(* Logix 5000 project; controller FV vendor 1 type 14 code 217 rev 31.11; software revision 31.00; part 38 of 63 *)
(* tags used below, declared in another part *)
   CWD : CHECKWORD_FLAGS;
   Dummy : BOOL;
   FV_Copy_from_fv_file : DINT;
   FV_Copy_to_fv_file : DINT;
   FV_LTX_YS_001 : PlantItem;   // LTX_YS_001
   FV_LTX_YS_001_RawInput : ALIAS FOR Remote_IO:7:I.Data.16;   // FV_LTX_YS_001
   FV_LTX_YS_002 : PlantItem;   // LTX_YS_002
   FV_LTX_YS_002_RawInput : ALIAS FOR Remote_IO:7:I.Data.17;   // FV_LTX_YS_002
   FV_N110 : INT[255];   // FV DATA 0 CURRENT FV DATA
   FV_N111 : INT[50];   // FV1, CURRENT FV DATA
   FV_N112 : INT[50];   // FV2, CURRENT FV DATA
   FV_N113 : INT[50];   // FV3, CURRENT FV DATA
   FV_N114 : INT[50];   // FV4, CURRENT FV DATA
   FV_N115 : INT[50];   // FV5, CURRENT FV DATA
   FV_N116 : INT[50];   // FV6, CURRENT FV DATA
   FV_N117 : INT[50];   // FV7, CURRENT FV DATA
   FV_N118 : INT[50];   // FV8, CURRENT FV DATA
   FV_N119 : INT[50];   // FV9, CURRENT FV DATA
   FV_N120 : INT[50];   // FV10, CURRENT FV DATA
   FV_N121 : INT[50];   // FV11, CURRENT FV DATA
   FV_N122 : INT[50];   // FV12, CURRENT FV DATA
   FV_N123 : INT[50];   // FV13, CURRENT FV DATA
   FV_N124 : INT[50];   // FV14, CURRENT FV DATA
   FV_N125 : INT[50];   // FV15, CURRENT FV DATA
   FV_N126 : INT[50];   // FV16, CURRENT FV DATA
   FV_N127 : INT[50];   // FV17, CURRENT FV DATA
   FV_N128 : INT[50];   // FV18, CURRENT FV DATA
   FV_N129 : INT[50];   // FV19, CURRENT FV DATA
   FV_N130 : INT[50];   // FV20, CURRENT FV DATA
   FV_N131 : INT[50];   // FV21, CURRENT FV DATA
   FV_N132 : INT[50];   // FV22, CURRENT FV DATA
   FV_N133 : INT[50];   // FV23, CURRENT FV DATA
   FV_N134 : INT[50];   // FV24, CURRENT FV DATA
   FV_N135 : INT[50];   // FV25, CURRENT FV DATA
   FV_N136 : INT[50];   // YSV1, CURRENT FV DATA
   FV_N137 : INT[50];   // YSV2, CURRENT FV DATA
   FV_N138 : INT[50];   // YSV3, CURRENT FV DATA
   FV_N139 : INT[255];   // YST1
   FV_N140 : INT[255];   // YST2
   FV_N141 : INT[255];   // YSV1 DATA
   FV_N142 : INT[255];   // YSV2 DATA
   FV_N143 : INT[255];   // YSV3 DATA
   FV_N144 : INT[255];   // YST1 DATA
   FV_N145 : INT[255];   // YST2 DATA
   FV_N146 : INT[50];   // FV26, CURRENT FV DATA
   FV_N147 : INT[50];   // FV27, CURRENT FV DATA
   FV_N148 : INT[50];   // FV28, CURRENT FV DATA
   FV_N149 : INT[50];   // FV29, CURRENT FV DATA
   FV_N150 : INT[50];   // FV30, CURRENT FV DATA
   FV_N151 : INT[50];   // FV31, CURRENT FV DATA
   FV_PX1 : PlantItem;   // PX1
   FV_PX1_RawInput : ALIAS FOR Remote_IO:6:I.Data.13;   // FV_PX1 Water flush proxy switch
   FV_PX2 : PlantItem;   // PX2
   FV_PX2_RawInput : ALIAS FOR Remote_IO:6:I.Data.14;   // FV_PX2 CIP supply proxy switch
   FV_PX3 : PlantItem;   // PX3
   FV_PX3_RawInput : ALIAS FOR Remote_IO:6:I.Data.15;   // FV_PX3 YSV1 to reseeding main proxy switch
   One_Second_One_Scan : ALIAS FOR One_Second_1_scan;
(* FV_Common, continued *)

ROUTINE FV_Copy_Vessel_File   (* ladder *)
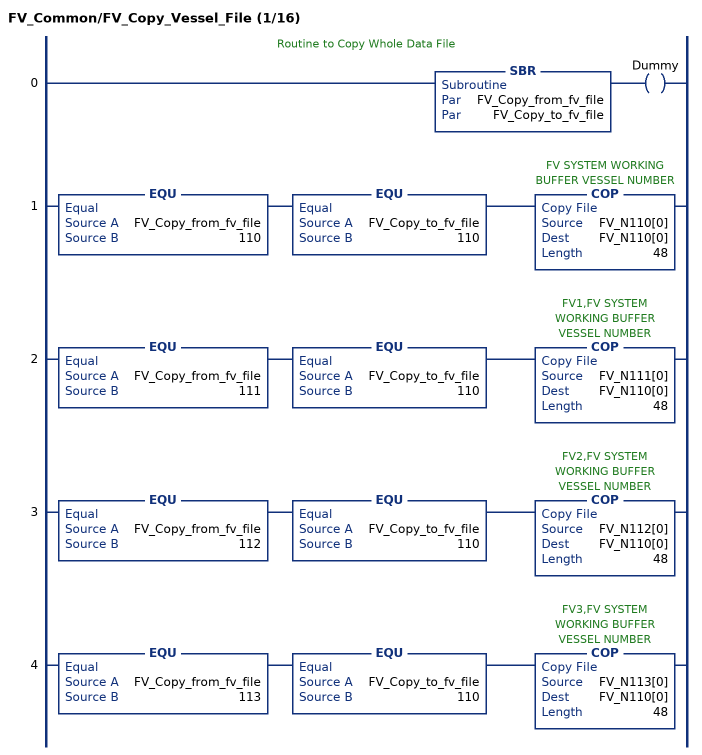
   // Routine to Copy Whole Data File
   0: SBR(FV_Copy_from_fv_file,FV_Copy_to_fv_file)OTE(Dummy);
   1: EQU(FV_Copy_from_fv_file,110)EQU(FV_Copy_to_fv_file,110)COP(FV_N110[0],FV_N110[0],48);
   2: EQU(FV_Copy_from_fv_file,111)EQU(FV_Copy_to_fv_file,110)COP(FV_N111[0],FV_N110[0],48);
   3: EQU(FV_Copy_from_fv_file,112)EQU(FV_Copy_to_fv_file,110)COP(FV_N112[0],FV_N110[0],48);
   4: EQU(FV_Copy_from_fv_file,113)EQU(FV_Copy_to_fv_file,110)COP(FV_N113[0],FV_N110[0],48);
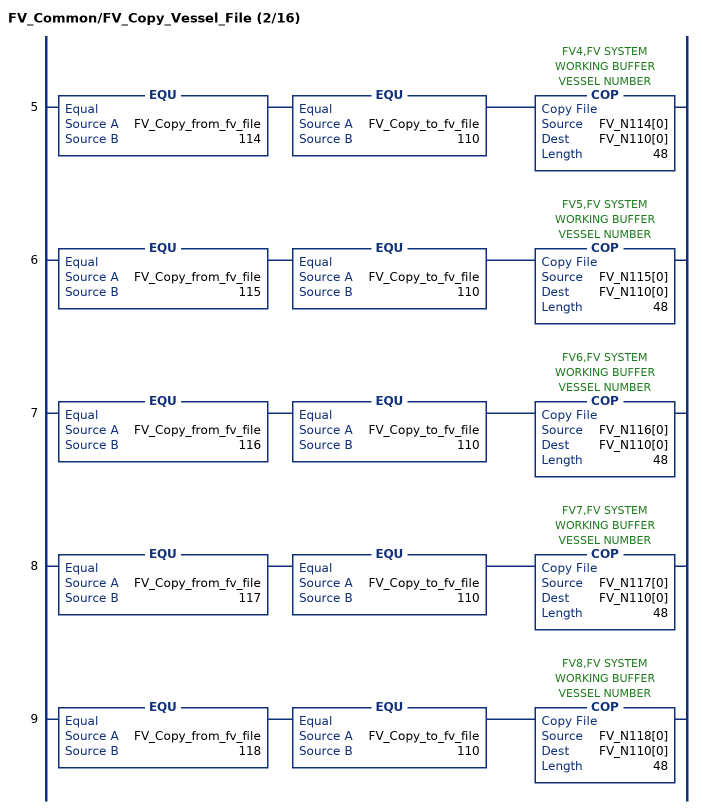
   5: EQU(FV_Copy_from_fv_file,114)EQU(FV_Copy_to_fv_file,110)COP(FV_N114[0],FV_N110[0],48);
   6: EQU(FV_Copy_from_fv_file,115)EQU(FV_Copy_to_fv_file,110)COP(FV_N115[0],FV_N110[0],48);
   7: EQU(FV_Copy_from_fv_file,116)EQU(FV_Copy_to_fv_file,110)COP(FV_N116[0],FV_N110[0],48);
   8: EQU(FV_Copy_from_fv_file,117)EQU(FV_Copy_to_fv_file,110)COP(FV_N117[0],FV_N110[0],48);
   9: EQU(FV_Copy_from_fv_file,118)EQU(FV_Copy_to_fv_file,110)COP(FV_N118[0],FV_N110[0],48);
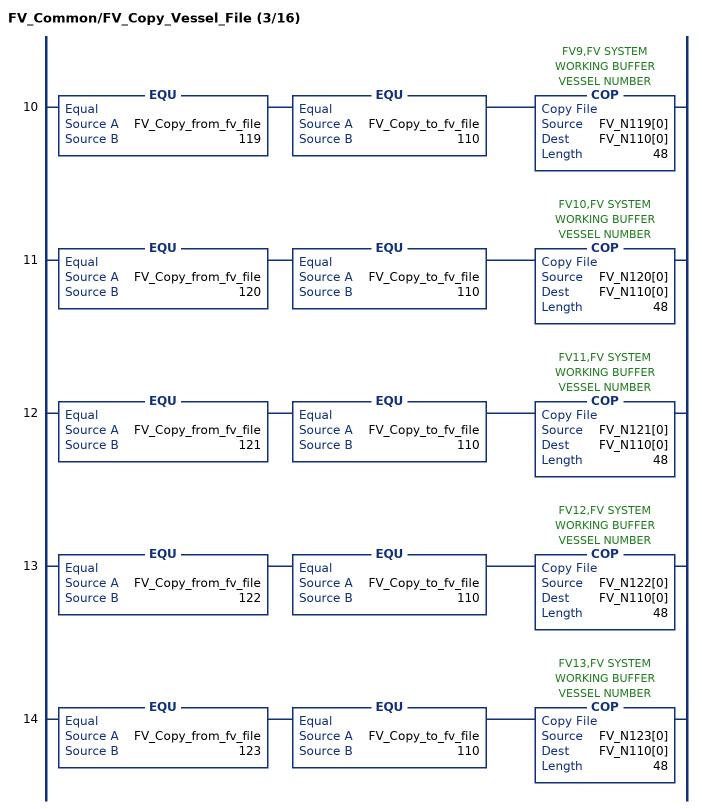
   10: EQU(FV_Copy_from_fv_file,119)EQU(FV_Copy_to_fv_file,110)COP(FV_N119[0],FV_N110[0],48);
   11: EQU(FV_Copy_from_fv_file,120)EQU(FV_Copy_to_fv_file,110)COP(FV_N120[0],FV_N110[0],48);
   12: EQU(FV_Copy_from_fv_file,121)EQU(FV_Copy_to_fv_file,110)COP(FV_N121[0],FV_N110[0],48);
   13: EQU(FV_Copy_from_fv_file,122)EQU(FV_Copy_to_fv_file,110)COP(FV_N122[0],FV_N110[0],48);
   14: EQU(FV_Copy_from_fv_file,123)EQU(FV_Copy_to_fv_file,110)COP(FV_N123[0],FV_N110[0],48);
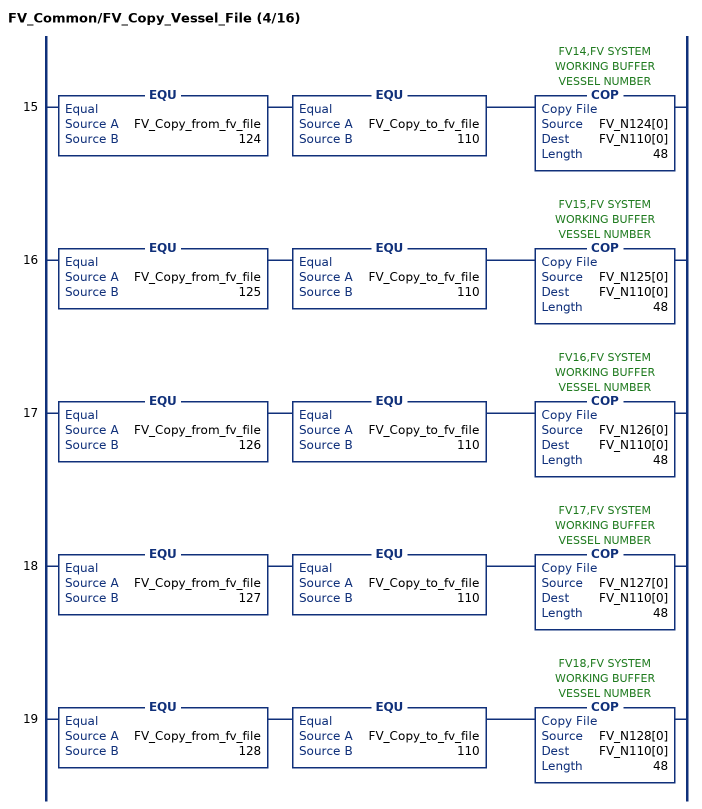
   15: EQU(FV_Copy_from_fv_file,124)EQU(FV_Copy_to_fv_file,110)COP(FV_N124[0],FV_N110[0],48);
   16: EQU(FV_Copy_from_fv_file,125)EQU(FV_Copy_to_fv_file,110)COP(FV_N125[0],FV_N110[0],48);
   17: EQU(FV_Copy_from_fv_file,126)EQU(FV_Copy_to_fv_file,110)COP(FV_N126[0],FV_N110[0],48);
   18: EQU(FV_Copy_from_fv_file,127)EQU(FV_Copy_to_fv_file,110)COP(FV_N127[0],FV_N110[0],48);
   19: EQU(FV_Copy_from_fv_file,128)EQU(FV_Copy_to_fv_file,110)COP(FV_N128[0],FV_N110[0],48);
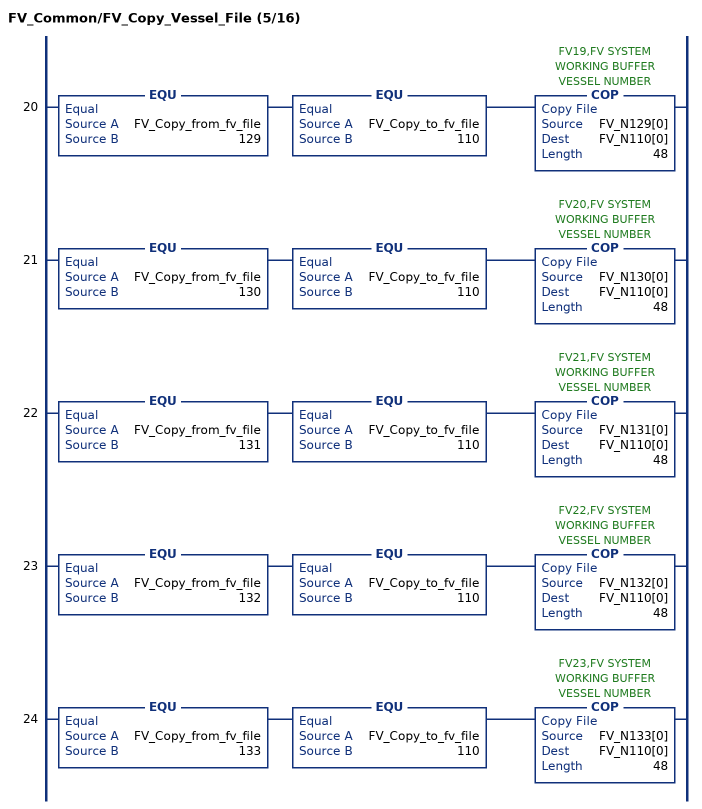
   20: EQU(FV_Copy_from_fv_file,129)EQU(FV_Copy_to_fv_file,110)COP(FV_N129[0],FV_N110[0],48);
   21: EQU(FV_Copy_from_fv_file,130)EQU(FV_Copy_to_fv_file,110)COP(FV_N130[0],FV_N110[0],48);
   22: EQU(FV_Copy_from_fv_file,131)EQU(FV_Copy_to_fv_file,110)COP(FV_N131[0],FV_N110[0],48);
   23: EQU(FV_Copy_from_fv_file,132)EQU(FV_Copy_to_fv_file,110)COP(FV_N132[0],FV_N110[0],48);
   24: EQU(FV_Copy_from_fv_file,133)EQU(FV_Copy_to_fv_file,110)COP(FV_N133[0],FV_N110[0],48);
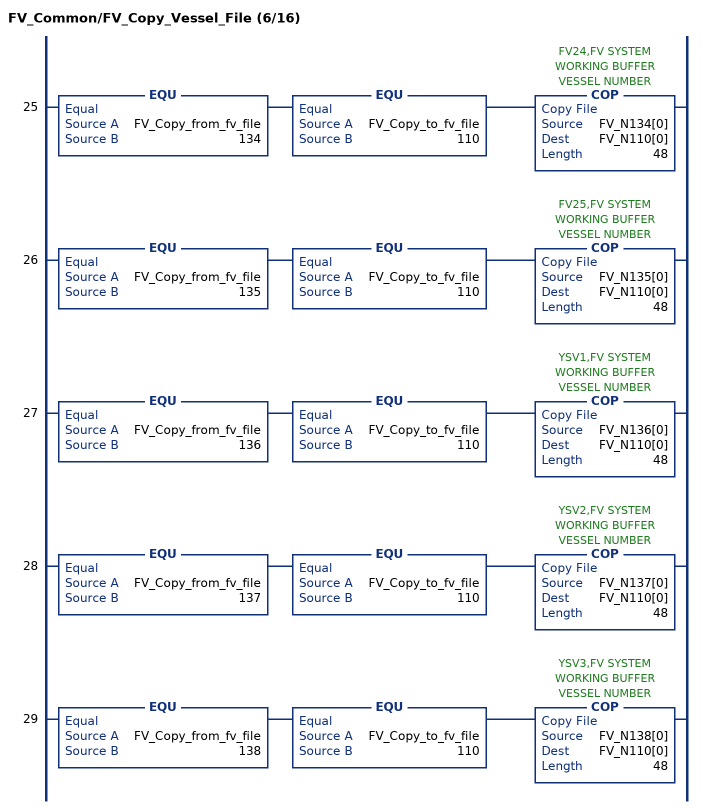
   25: EQU(FV_Copy_from_fv_file,134)EQU(FV_Copy_to_fv_file,110)COP(FV_N134[0],FV_N110[0],48);
   26: EQU(FV_Copy_from_fv_file,135)EQU(FV_Copy_to_fv_file,110)COP(FV_N135[0],FV_N110[0],48);
   27: EQU(FV_Copy_from_fv_file,136)EQU(FV_Copy_to_fv_file,110)COP(FV_N136[0],FV_N110[0],48);
   28: EQU(FV_Copy_from_fv_file,137)EQU(FV_Copy_to_fv_file,110)COP(FV_N137[0],FV_N110[0],48);
   29: EQU(FV_Copy_from_fv_file,138)EQU(FV_Copy_to_fv_file,110)COP(FV_N138[0],FV_N110[0],48);
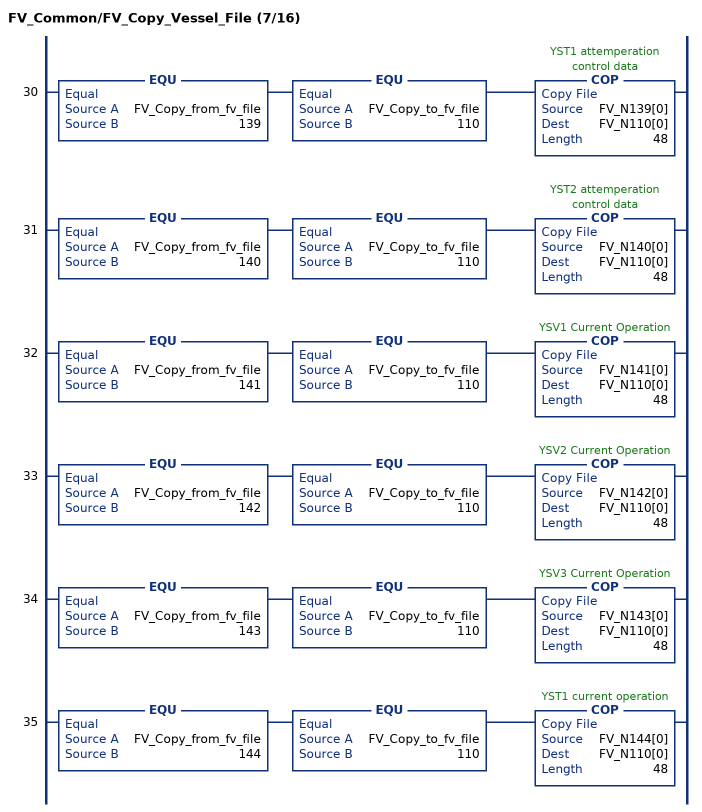
   30: EQU(FV_Copy_from_fv_file,139)EQU(FV_Copy_to_fv_file,110)COP(FV_N139[0],FV_N110[0],48);
   31: EQU(FV_Copy_from_fv_file,140)EQU(FV_Copy_to_fv_file,110)COP(FV_N140[0],FV_N110[0],48);
   32: EQU(FV_Copy_from_fv_file,141)EQU(FV_Copy_to_fv_file,110)COP(FV_N141[0],FV_N110[0],48);
   33: EQU(FV_Copy_from_fv_file,142)EQU(FV_Copy_to_fv_file,110)COP(FV_N142[0],FV_N110[0],48);
   34: EQU(FV_Copy_from_fv_file,143)EQU(FV_Copy_to_fv_file,110)COP(FV_N143[0],FV_N110[0],48);
   35: EQU(FV_Copy_from_fv_file,144)EQU(FV_Copy_to_fv_file,110)COP(FV_N144[0],FV_N110[0],48);
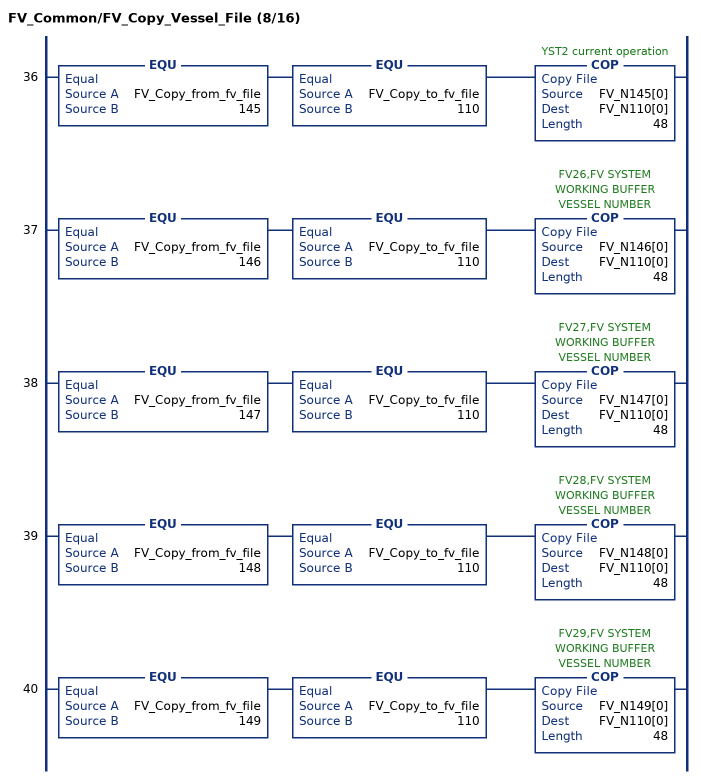
   36: EQU(FV_Copy_from_fv_file,145)EQU(FV_Copy_to_fv_file,110)COP(FV_N145[0],FV_N110[0],48);
   37: EQU(FV_Copy_from_fv_file,146)EQU(FV_Copy_to_fv_file,110)COP(FV_N146[0],FV_N110[0],48);
   38: EQU(FV_Copy_from_fv_file,147)EQU(FV_Copy_to_fv_file,110)COP(FV_N147[0],FV_N110[0],48);
   39: EQU(FV_Copy_from_fv_file,148)EQU(FV_Copy_to_fv_file,110)COP(FV_N148[0],FV_N110[0],48);
   40: EQU(FV_Copy_from_fv_file,149)EQU(FV_Copy_to_fv_file,110)COP(FV_N149[0],FV_N110[0],48);
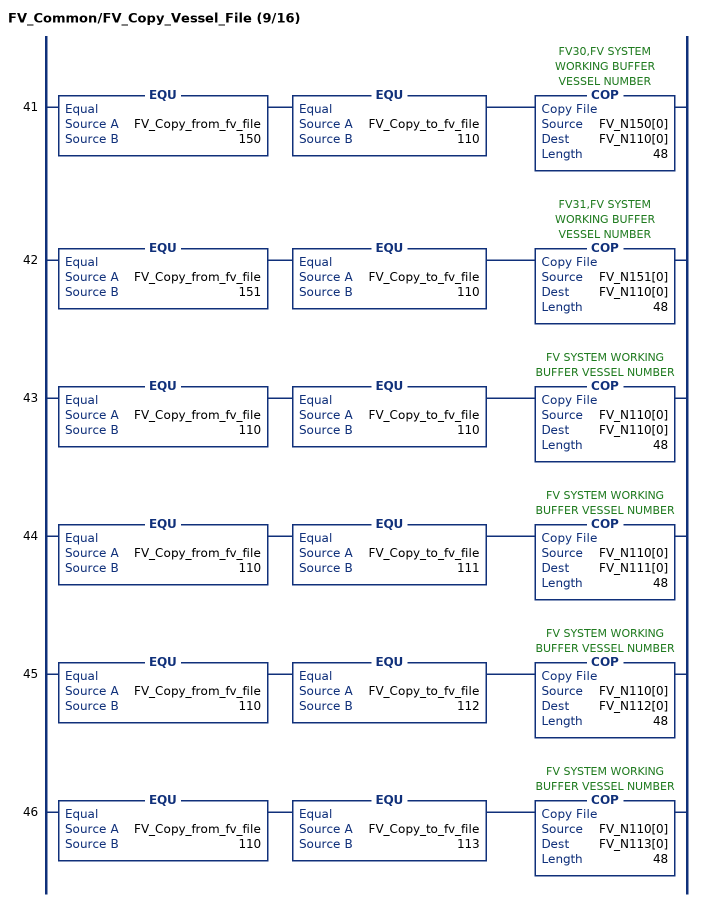
   41: EQU(FV_Copy_from_fv_file,150)EQU(FV_Copy_to_fv_file,110)COP(FV_N150[0],FV_N110[0],48);
   42: EQU(FV_Copy_from_fv_file,151)EQU(FV_Copy_to_fv_file,110)COP(FV_N151[0],FV_N110[0],48);
   43: EQU(FV_Copy_from_fv_file,110)EQU(FV_Copy_to_fv_file,110)COP(FV_N110[0],FV_N110[0],48);
   44: EQU(FV_Copy_from_fv_file,110)EQU(FV_Copy_to_fv_file,111)COP(FV_N110[0],FV_N111[0],48);
   45: EQU(FV_Copy_from_fv_file,110)EQU(FV_Copy_to_fv_file,112)COP(FV_N110[0],FV_N112[0],48);
   46: EQU(FV_Copy_from_fv_file,110)EQU(FV_Copy_to_fv_file,113)COP(FV_N110[0],FV_N113[0],48);
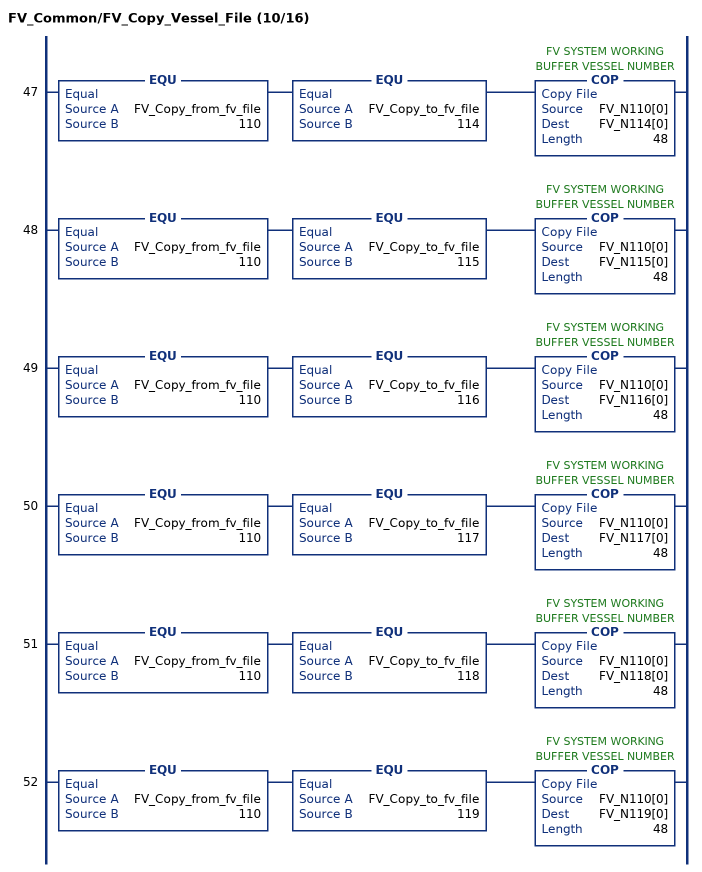
   47: EQU(FV_Copy_from_fv_file,110)EQU(FV_Copy_to_fv_file,114)COP(FV_N110[0],FV_N114[0],48);
   48: EQU(FV_Copy_from_fv_file,110)EQU(FV_Copy_to_fv_file,115)COP(FV_N110[0],FV_N115[0],48);
   49: EQU(FV_Copy_from_fv_file,110)EQU(FV_Copy_to_fv_file,116)COP(FV_N110[0],FV_N116[0],48);
   50: EQU(FV_Copy_from_fv_file,110)EQU(FV_Copy_to_fv_file,117)COP(FV_N110[0],FV_N117[0],48);
   51: EQU(FV_Copy_from_fv_file,110)EQU(FV_Copy_to_fv_file,118)COP(FV_N110[0],FV_N118[0],48);
   52: EQU(FV_Copy_from_fv_file,110)EQU(FV_Copy_to_fv_file,119)COP(FV_N110[0],FV_N119[0],48);
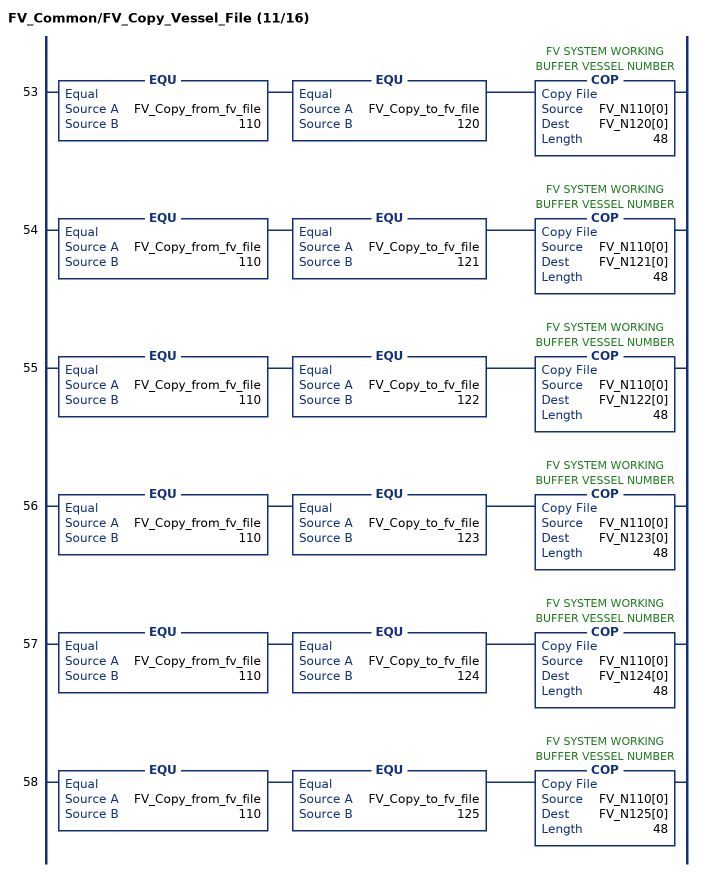
   53: EQU(FV_Copy_from_fv_file,110)EQU(FV_Copy_to_fv_file,120)COP(FV_N110[0],FV_N120[0],48);
   54: EQU(FV_Copy_from_fv_file,110)EQU(FV_Copy_to_fv_file,121)COP(FV_N110[0],FV_N121[0],48);
   55: EQU(FV_Copy_from_fv_file,110)EQU(FV_Copy_to_fv_file,122)COP(FV_N110[0],FV_N122[0],48);
   56: EQU(FV_Copy_from_fv_file,110)EQU(FV_Copy_to_fv_file,123)COP(FV_N110[0],FV_N123[0],48);
   57: EQU(FV_Copy_from_fv_file,110)EQU(FV_Copy_to_fv_file,124)COP(FV_N110[0],FV_N124[0],48);
   58: EQU(FV_Copy_from_fv_file,110)EQU(FV_Copy_to_fv_file,125)COP(FV_N110[0],FV_N125[0],48);
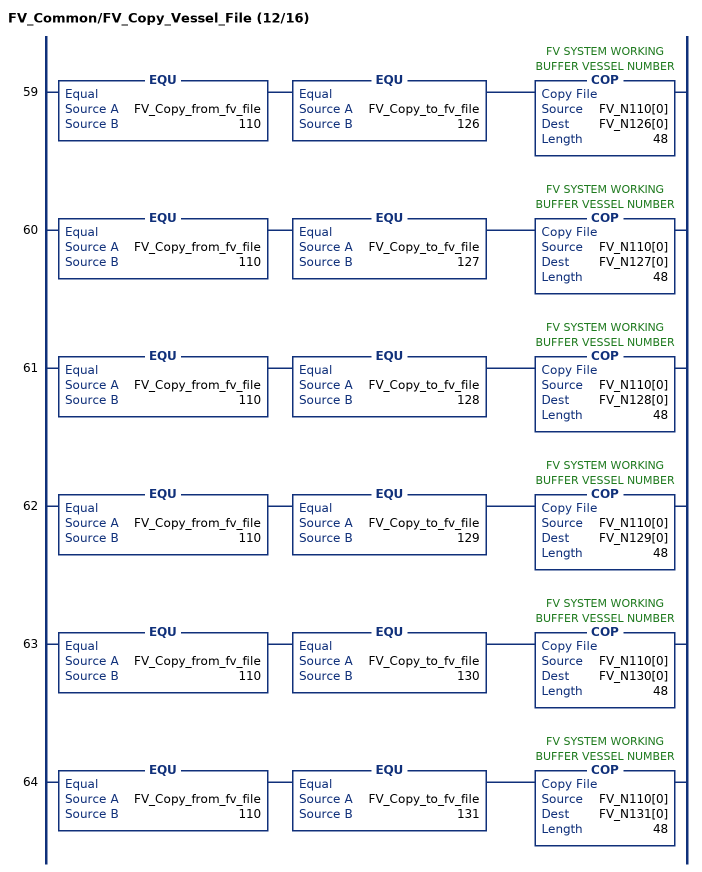
   59: EQU(FV_Copy_from_fv_file,110)EQU(FV_Copy_to_fv_file,126)COP(FV_N110[0],FV_N126[0],48);
   60: EQU(FV_Copy_from_fv_file,110)EQU(FV_Copy_to_fv_file,127)COP(FV_N110[0],FV_N127[0],48);
   61: EQU(FV_Copy_from_fv_file,110)EQU(FV_Copy_to_fv_file,128)COP(FV_N110[0],FV_N128[0],48);
   62: EQU(FV_Copy_from_fv_file,110)EQU(FV_Copy_to_fv_file,129)COP(FV_N110[0],FV_N129[0],48);
   63: EQU(FV_Copy_from_fv_file,110)EQU(FV_Copy_to_fv_file,130)COP(FV_N110[0],FV_N130[0],48);
   64: EQU(FV_Copy_from_fv_file,110)EQU(FV_Copy_to_fv_file,131)COP(FV_N110[0],FV_N131[0],48);
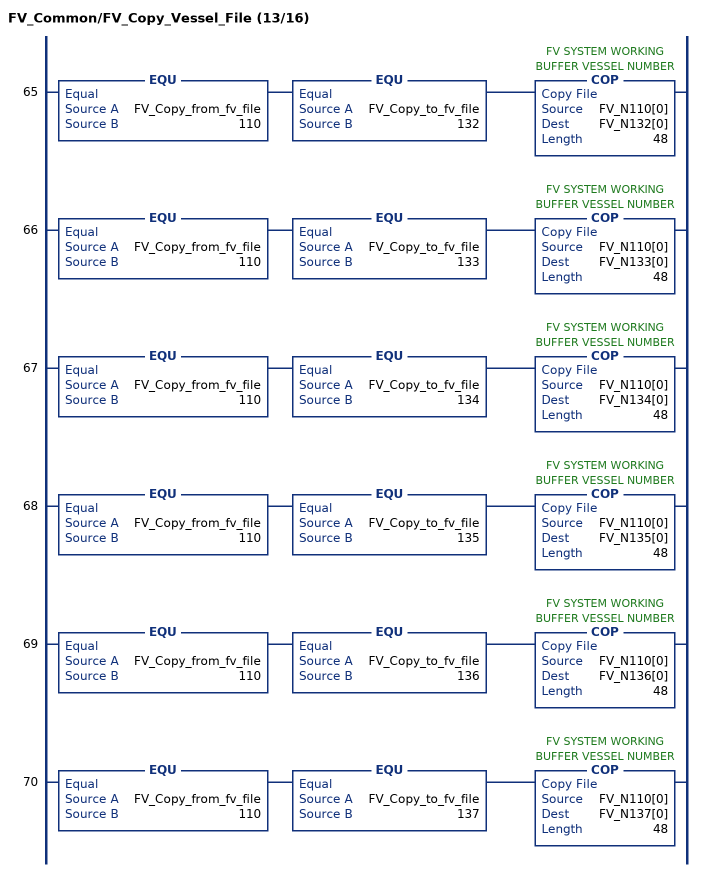
   65: EQU(FV_Copy_from_fv_file,110)EQU(FV_Copy_to_fv_file,132)COP(FV_N110[0],FV_N132[0],48);
   66: EQU(FV_Copy_from_fv_file,110)EQU(FV_Copy_to_fv_file,133)COP(FV_N110[0],FV_N133[0],48);
   67: EQU(FV_Copy_from_fv_file,110)EQU(FV_Copy_to_fv_file,134)COP(FV_N110[0],FV_N134[0],48);
   68: EQU(FV_Copy_from_fv_file,110)EQU(FV_Copy_to_fv_file,135)COP(FV_N110[0],FV_N135[0],48);
   69: EQU(FV_Copy_from_fv_file,110)EQU(FV_Copy_to_fv_file,136)COP(FV_N110[0],FV_N136[0],48);
   70: EQU(FV_Copy_from_fv_file,110)EQU(FV_Copy_to_fv_file,137)COP(FV_N110[0],FV_N137[0],48);
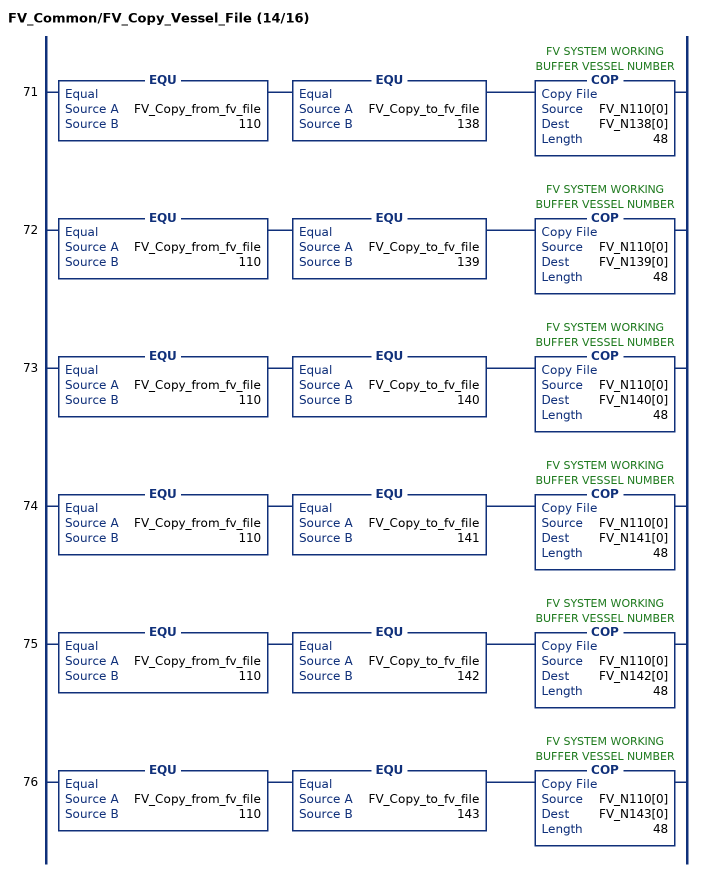
   71: EQU(FV_Copy_from_fv_file,110)EQU(FV_Copy_to_fv_file,138)COP(FV_N110[0],FV_N138[0],48);
   72: EQU(FV_Copy_from_fv_file,110)EQU(FV_Copy_to_fv_file,139)COP(FV_N110[0],FV_N139[0],48);
   73: EQU(FV_Copy_from_fv_file,110)EQU(FV_Copy_to_fv_file,140)COP(FV_N110[0],FV_N140[0],48);
   74: EQU(FV_Copy_from_fv_file,110)EQU(FV_Copy_to_fv_file,141)COP(FV_N110[0],FV_N141[0],48);
   75: EQU(FV_Copy_from_fv_file,110)EQU(FV_Copy_to_fv_file,142)COP(FV_N110[0],FV_N142[0],48);
   76: EQU(FV_Copy_from_fv_file,110)EQU(FV_Copy_to_fv_file,143)COP(FV_N110[0],FV_N143[0],48);
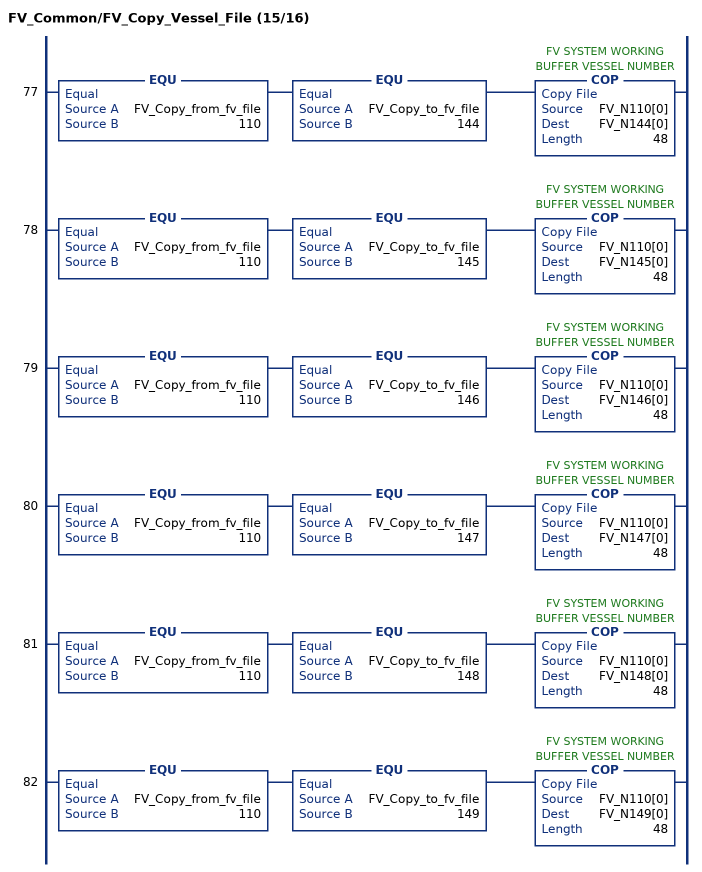
   77: EQU(FV_Copy_from_fv_file,110)EQU(FV_Copy_to_fv_file,144)COP(FV_N110[0],FV_N144[0],48);
   78: EQU(FV_Copy_from_fv_file,110)EQU(FV_Copy_to_fv_file,145)COP(FV_N110[0],FV_N145[0],48);
   79: EQU(FV_Copy_from_fv_file,110)EQU(FV_Copy_to_fv_file,146)COP(FV_N110[0],FV_N146[0],48);
   80: EQU(FV_Copy_from_fv_file,110)EQU(FV_Copy_to_fv_file,147)COP(FV_N110[0],FV_N147[0],48);
   81: EQU(FV_Copy_from_fv_file,110)EQU(FV_Copy_to_fv_file,148)COP(FV_N110[0],FV_N148[0],48);
   82: EQU(FV_Copy_from_fv_file,110)EQU(FV_Copy_to_fv_file,149)COP(FV_N110[0],FV_N149[0],48);
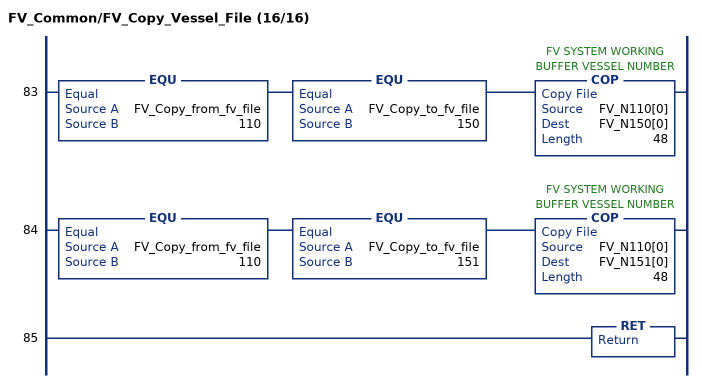
   83: EQU(FV_Copy_from_fv_file,110)EQU(FV_Copy_to_fv_file,150)COP(FV_N110[0],FV_N150[0],48);
   84: EQU(FV_Copy_from_fv_file,110)EQU(FV_Copy_to_fv_file,151)COP(FV_N110[0],FV_N151[0],48);
   85: RET();
END_ROUTINE

ROUTINE FV_DEBOUNCE_8   (* ladder *)
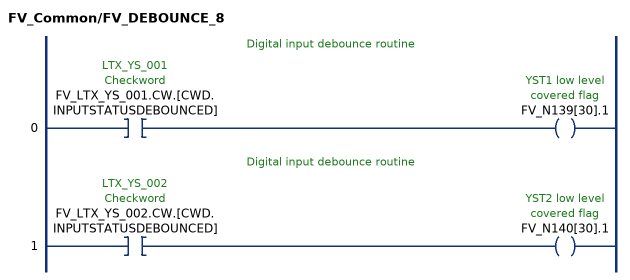
   // Digital input debounce routine
   0: XIC(FV_LTX_YS_001.CW.[CWD.INPUTSTATUSDEBOUNCED])OTE(FV_N139[30].1);
   // Digital input debounce routine
   1: XIC(FV_LTX_YS_002.CW.[CWD.INPUTSTATUSDEBOUNCED])OTE(FV_N140[30].1);
END_ROUTINE

ROUTINE FV_Digital_Inputs   (* ladder *)
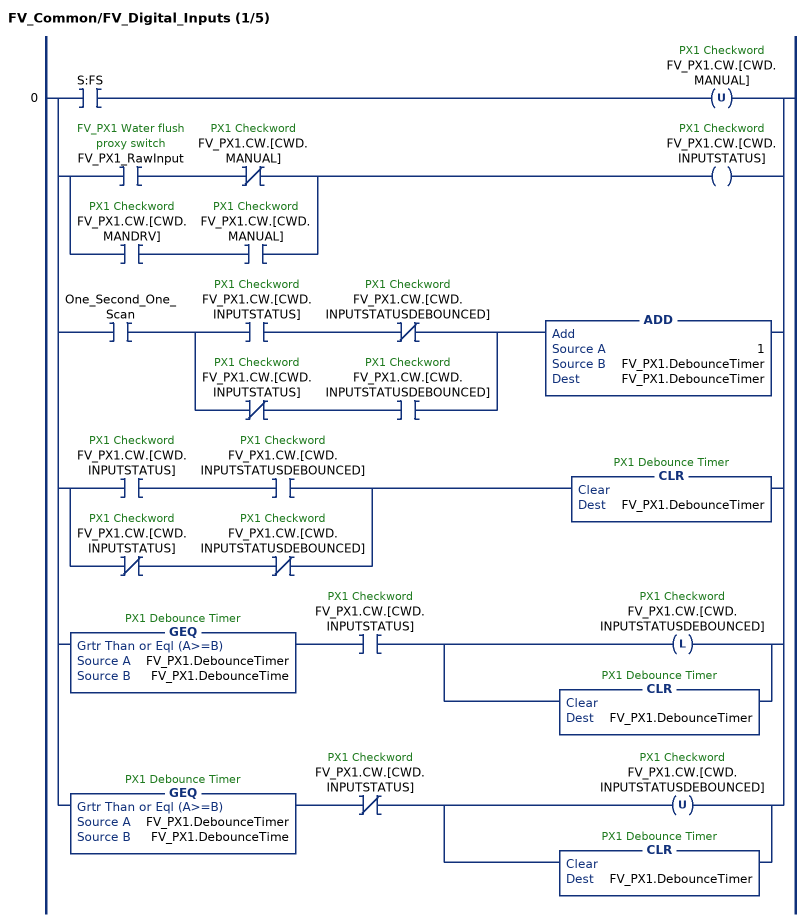
   0: [XIC(S:FS) OTU(FV_PX1.CW.[CWD.MANUAL]) ,[XIC(FV_PX1_RawInput) XIO(FV_PX1.CW.[CWD.MANUAL]) ,XIC(FV_PX1.CW.[CWD.MANDRV]) XIC(FV_PX1.CW.[CWD.MANUAL]) ] OTE(FV_PX1.CW.[CWD.INPUTSTATUS]) ,XIC(One_Second_One_Scan) [XIC(FV_PX1.CW.[CWD.INPUTSTATUS]) XIO(FV_PX1.CW.[CWD.INPUTSTATUSDEBOUNCED]) ,XIO(FV_PX1.CW.[CWD.INPUTSTATUS]) XIC(FV_PX1.CW.[CWD.INPUTSTATUSDEBOUNCED]) ] ADD(1,FV_PX1.DebounceTimer,FV_PX1.DebounceTimer) ,[XIC(FV_PX1.CW.[CWD.INPUTSTATUS]) XIC(FV_PX1.CW.[CWD.INPUTSTATUSDEBOUNCED]) ,XIO(FV_PX1.CW.[CWD.INPUTSTATUS]) XIO(FV_PX1.CW.[CWD.INPUTSTATUSDEBOUNCED]) ] CLR(FV_PX1.DebounceTimer) ,GEQ(FV_PX1.DebounceTimer,FV_PX1.DebounceTime) XIC(FV_PX1.CW.[CWD.INPUTSTATUS]) [OTL(FV_PX1.CW.[CWD.INPUTSTATUSDEBOUNCED]) ,CLR(FV_PX1.DebounceTimer) ] ,GEQ(FV_PX1.DebounceTimer,FV_PX1.DebounceTime) XIO(FV_PX1.CW.[CWD.INPUTSTATUS]) [OTU(FV_PX1.CW.[CWD.INPUTSTATUSDEBOUNCED]) ,CLR(FV_PX1.DebounceTimer) ] ];
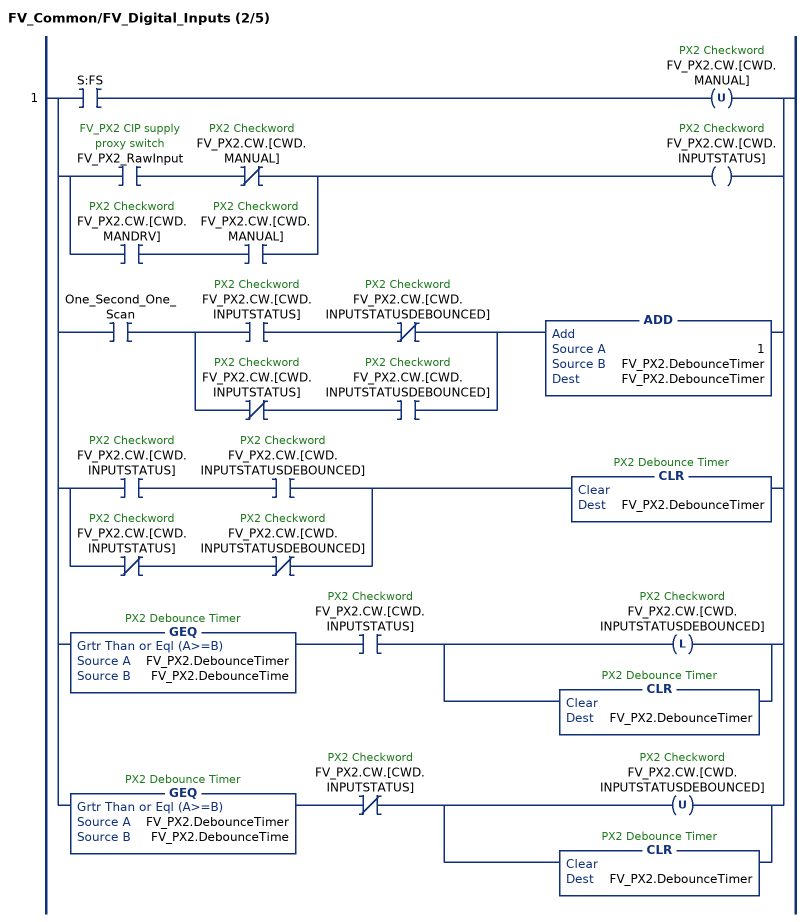
   1: [XIC(S:FS) OTU(FV_PX2.CW.[CWD.MANUAL]) ,[XIC(FV_PX2_RawInput) XIO(FV_PX2.CW.[CWD.MANUAL]) ,XIC(FV_PX2.CW.[CWD.MANDRV]) XIC(FV_PX2.CW.[CWD.MANUAL]) ] OTE(FV_PX2.CW.[CWD.INPUTSTATUS]) ,XIC(One_Second_One_Scan) [XIC(FV_PX2.CW.[CWD.INPUTSTATUS]) XIO(FV_PX2.CW.[CWD.INPUTSTATUSDEBOUNCED]) ,XIO(FV_PX2.CW.[CWD.INPUTSTATUS]) XIC(FV_PX2.CW.[CWD.INPUTSTATUSDEBOUNCED]) ] ADD(1,FV_PX2.DebounceTimer,FV_PX2.DebounceTimer) ,[XIC(FV_PX2.CW.[CWD.INPUTSTATUS]) XIC(FV_PX2.CW.[CWD.INPUTSTATUSDEBOUNCED]) ,XIO(FV_PX2.CW.[CWD.INPUTSTATUS]) XIO(FV_PX2.CW.[CWD.INPUTSTATUSDEBOUNCED]) ] CLR(FV_PX2.DebounceTimer) ,GEQ(FV_PX2.DebounceTimer,FV_PX2.DebounceTime) XIC(FV_PX2.CW.[CWD.INPUTSTATUS]) [OTL(FV_PX2.CW.[CWD.INPUTSTATUSDEBOUNCED]) ,CLR(FV_PX2.DebounceTimer) ] ,GEQ(FV_PX2.DebounceTimer,FV_PX2.DebounceTime) XIO(FV_PX2.CW.[CWD.INPUTSTATUS]) [OTU(FV_PX2.CW.[CWD.INPUTSTATUSDEBOUNCED]) ,CLR(FV_PX2.DebounceTimer) ] ];
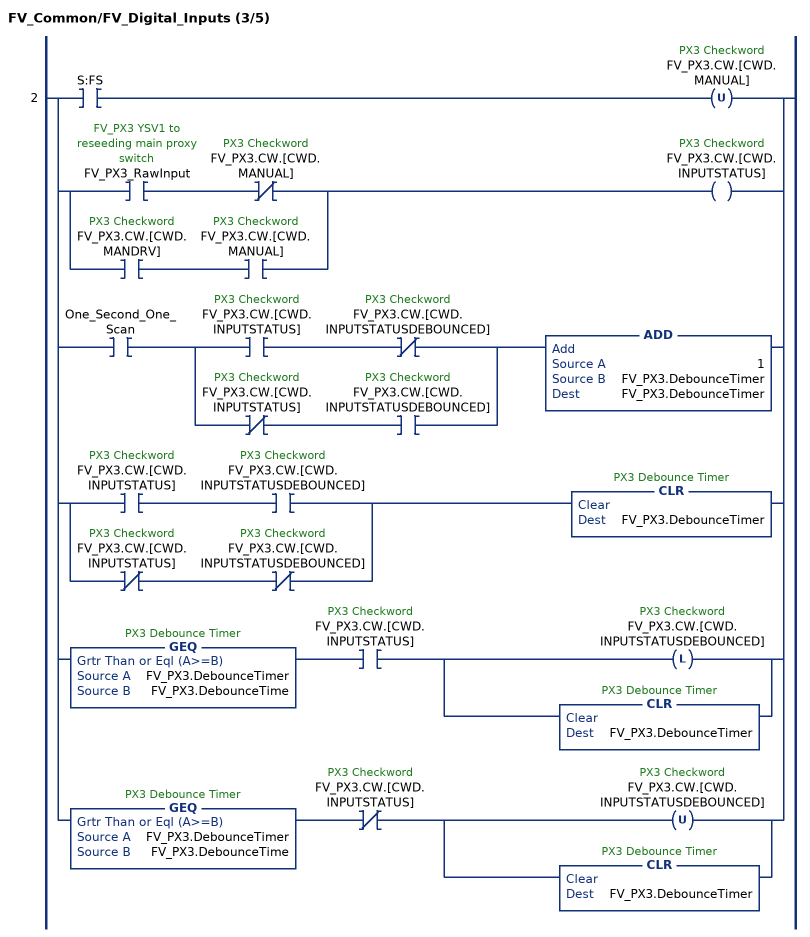
   2: [XIC(S:FS) OTU(FV_PX3.CW.[CWD.MANUAL]) ,[XIC(FV_PX3_RawInput) XIO(FV_PX3.CW.[CWD.MANUAL]) ,XIC(FV_PX3.CW.[CWD.MANDRV]) XIC(FV_PX3.CW.[CWD.MANUAL]) ] OTE(FV_PX3.CW.[CWD.INPUTSTATUS]) ,XIC(One_Second_One_Scan) [XIC(FV_PX3.CW.[CWD.INPUTSTATUS]) XIO(FV_PX3.CW.[CWD.INPUTSTATUSDEBOUNCED]) ,XIO(FV_PX3.CW.[CWD.INPUTSTATUS]) XIC(FV_PX3.CW.[CWD.INPUTSTATUSDEBOUNCED]) ] ADD(1,FV_PX3.DebounceTimer,FV_PX3.DebounceTimer) ,[XIC(FV_PX3.CW.[CWD.INPUTSTATUS]) XIC(FV_PX3.CW.[CWD.INPUTSTATUSDEBOUNCED]) ,XIO(FV_PX3.CW.[CWD.INPUTSTATUS]) XIO(FV_PX3.CW.[CWD.INPUTSTATUSDEBOUNCED]) ] CLR(FV_PX3.DebounceTimer) ,GEQ(FV_PX3.DebounceTimer,FV_PX3.DebounceTime) XIC(FV_PX3.CW.[CWD.INPUTSTATUS]) [OTL(FV_PX3.CW.[CWD.INPUTSTATUSDEBOUNCED]) ,CLR(FV_PX3.DebounceTimer) ] ,GEQ(FV_PX3.DebounceTimer,FV_PX3.DebounceTime) XIO(FV_PX3.CW.[CWD.INPUTSTATUS]) [OTU(FV_PX3.CW.[CWD.INPUTSTATUSDEBOUNCED]) ,CLR(FV_PX3.DebounceTimer) ] ];
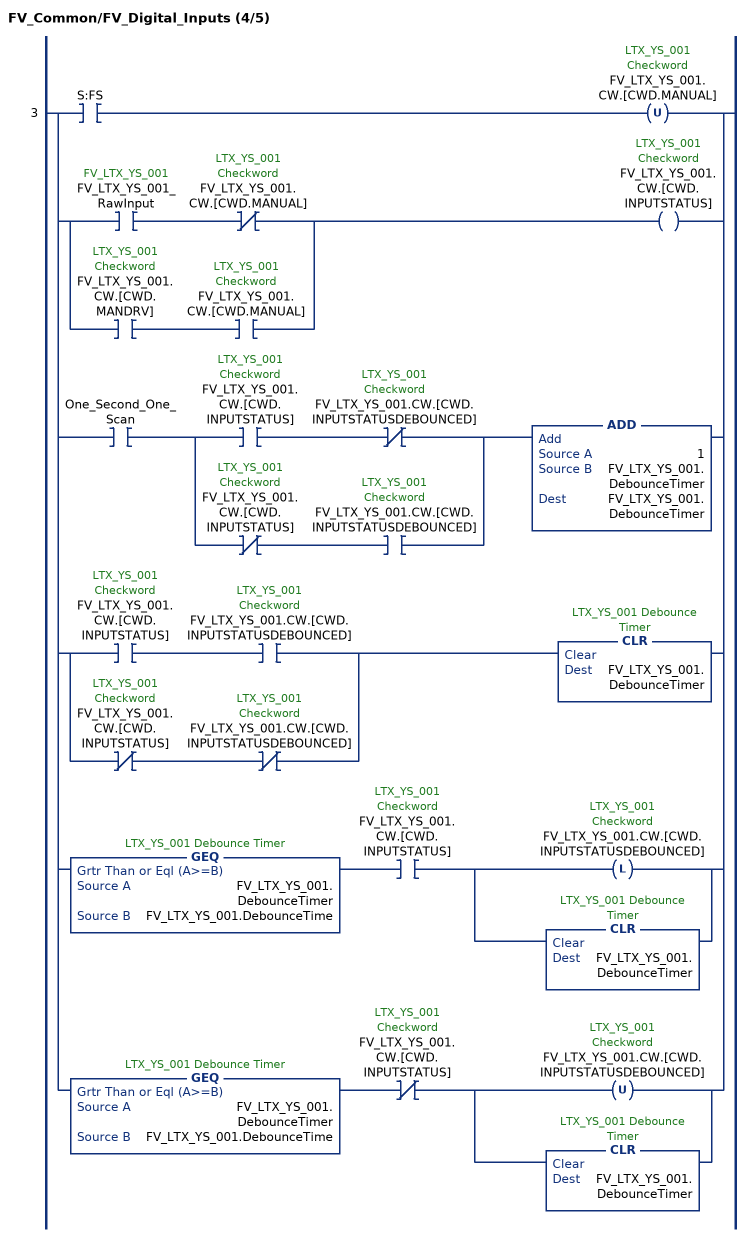
   3: [XIC(S:FS) OTU(FV_LTX_YS_001.CW.[CWD.MANUAL]) ,[XIC(FV_LTX_YS_001_RawInput) XIO(FV_LTX_YS_001.CW.[CWD.MANUAL]) ,XIC(FV_LTX_YS_001.CW.[CWD.MANDRV]) XIC(FV_LTX_YS_001.CW.[CWD.MANUAL]) ] OTE(FV_LTX_YS_001.CW.[CWD.INPUTSTATUS]) ,XIC(One_Second_One_Scan) [XIC(FV_LTX_YS_001.CW.[CWD.INPUTSTATUS]) XIO(FV_LTX_YS_001.CW.[CWD.INPUTSTATUSDEBOUNCED]) ,XIO(FV_LTX_YS_001.CW.[CWD.INPUTSTATUS]) XIC(FV_LTX_YS_001.CW.[CWD.INPUTSTATUSDEBOUNCED]) ] ADD(1,FV_LTX_YS_001.DebounceTimer,FV_LTX_YS_001.DebounceTimer) ,[XIC(FV_LTX_YS_001.CW.[CWD.INPUTSTATUS]) XIC(FV_LTX_YS_001.CW.[CWD.INPUTSTATUSDEBOUNCED]) ,XIO(FV_LTX_YS_001.CW.[CWD.INPUTSTATUS]) XIO(FV_LTX_YS_001.CW.[CWD.INPUTSTATUSDEBOUNCED]) ] CLR(FV_LTX_YS_001.DebounceTimer) ,GEQ(FV_LTX_YS_001.DebounceTimer,FV_LTX_YS_001.DebounceTime) XIC(FV_LTX_YS_001.CW.[CWD.INPUTSTATUS]) [OTL(FV_LTX_YS_001.CW.[CWD.INPUTSTATUSDEBOUNCED]) ,CLR(FV_LTX_YS_001.DebounceTimer) ] ,GEQ(FV_LTX_YS_001.DebounceTimer,FV_LTX_YS_001.DebounceTime) XIO(FV_LTX_YS_001.CW.[CWD.INPUTSTATUS]) [OTU(FV_LTX_YS_001.CW.[CWD.INPUTSTATUSDEBOUNCED]) ,CLR(FV_LTX_YS_001.DebounceTimer) ] ];
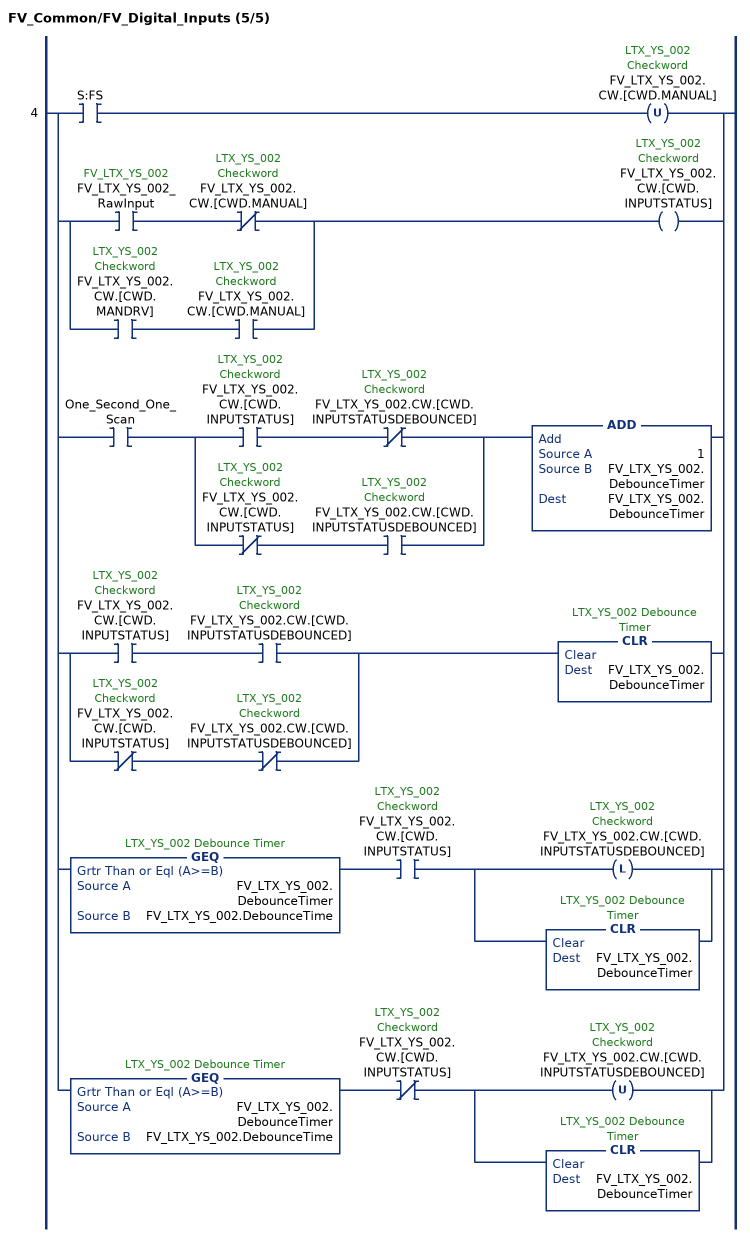
   4: [XIC(S:FS) OTU(FV_LTX_YS_002.CW.[CWD.MANUAL]) ,[XIC(FV_LTX_YS_002_RawInput) XIO(FV_LTX_YS_002.CW.[CWD.MANUAL]) ,XIC(FV_LTX_YS_002.CW.[CWD.MANDRV]) XIC(FV_LTX_YS_002.CW.[CWD.MANUAL]) ] OTE(FV_LTX_YS_002.CW.[CWD.INPUTSTATUS]) ,XIC(One_Second_One_Scan) [XIC(FV_LTX_YS_002.CW.[CWD.INPUTSTATUS]) XIO(FV_LTX_YS_002.CW.[CWD.INPUTSTATUSDEBOUNCED]) ,XIO(FV_LTX_YS_002.CW.[CWD.INPUTSTATUS]) XIC(FV_LTX_YS_002.CW.[CWD.INPUTSTATUSDEBOUNCED]) ] ADD(1,FV_LTX_YS_002.DebounceTimer,FV_LTX_YS_002.DebounceTimer) ,[XIC(FV_LTX_YS_002.CW.[CWD.INPUTSTATUS]) XIC(FV_LTX_YS_002.CW.[CWD.INPUTSTATUSDEBOUNCED]) ,XIO(FV_LTX_YS_002.CW.[CWD.INPUTSTATUS]) XIO(FV_LTX_YS_002.CW.[CWD.INPUTSTATUSDEBOUNCED]) ] CLR(FV_LTX_YS_002.DebounceTimer) ,GEQ(FV_LTX_YS_002.DebounceTimer,FV_LTX_YS_002.DebounceTime) XIC(FV_LTX_YS_002.CW.[CWD.INPUTSTATUS]) [OTL(FV_LTX_YS_002.CW.[CWD.INPUTSTATUSDEBOUNCED]) ,CLR(FV_LTX_YS_002.DebounceTimer) ] ,GEQ(FV_LTX_YS_002.DebounceTimer,FV_LTX_YS_002.DebounceTime) XIO(FV_LTX_YS_002.CW.[CWD.INPUTSTATUS]) [OTU(FV_LTX_YS_002.CW.[CWD.INPUTSTATUSDEBOUNCED]) ,CLR(FV_LTX_YS_002.DebounceTimer) ] ];
END_ROUTINE
